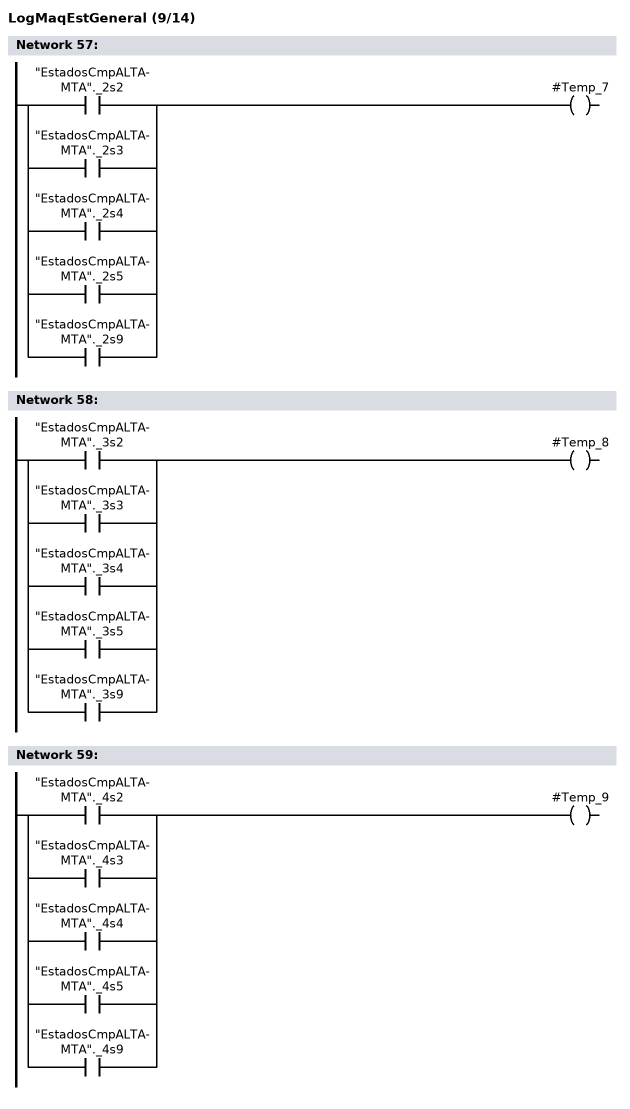
   RUNG wire#powerrail
      Contact( "EstadosCmpALTA-MTA"._2s2 )
      wire#w1
      Coil( #Temp_7 )
   END_RUNG
   RUNG wire#powerrail
      Contact( "EstadosCmpALTA-MTA"._2s3 )
   END_RUNG wire#w1
   RUNG wire#powerrail
      Contact( "EstadosCmpALTA-MTA"._2s4 )
   END_RUNG wire#w1
   RUNG wire#powerrail
      Contact( "EstadosCmpALTA-MTA"._2s5 )
   END_RUNG wire#w1
   RUNG wire#powerrail
      Contact( "EstadosCmpALTA-MTA"._2s9 )
   END_RUNG wire#w1
   // the same network as SCL:
   #Temp_7 := "EstadosCmpALTA-MTA"._2s2 OR "EstadosCmpALTA-MTA"._2s3 OR "EstadosCmpALTA-MTA"._2s4 OR "EstadosCmpALTA-MTA"._2s5 OR "EstadosCmpALTA-MTA"._2s9;
END_REGION

REGION Network 58
   RUNG wire#powerrail
      Contact( "EstadosCmpALTA-MTA"._3s2 )
      wire#w1
      Coil( #Temp_8 )
   END_RUNG
   RUNG wire#powerrail
      Contact( "EstadosCmpALTA-MTA"._3s3 )
   END_RUNG wire#w1
   RUNG wire#powerrail
      Contact( "EstadosCmpALTA-MTA"._3s4 )
   END_RUNG wire#w1
   RUNG wire#powerrail
      Contact( "EstadosCmpALTA-MTA"._3s5 )
   END_RUNG wire#w1
   RUNG wire#powerrail
      Contact( "EstadosCmpALTA-MTA"._3s9 )
   END_RUNG wire#w1
   // the same network as SCL:
   #Temp_8 := "EstadosCmpALTA-MTA"._3s2 OR "EstadosCmpALTA-MTA"._3s3 OR "EstadosCmpALTA-MTA"._3s4 OR "EstadosCmpALTA-MTA"._3s5 OR "EstadosCmpALTA-MTA"._3s9;
END_REGION

REGION Network 59
   RUNG wire#powerrail
      Contact( "EstadosCmpALTA-MTA"._4s2 )
      wire#w1
      Coil( #Temp_9 )
   END_RUNG
   RUNG wire#powerrail
      Contact( "EstadosCmpALTA-MTA"._4s3 )
   END_RUNG wire#w1
   RUNG wire#powerrail
      Contact( "EstadosCmpALTA-MTA"._4s4 )
   END_RUNG wire#w1
   RUNG wire#powerrail
      Contact( "EstadosCmpALTA-MTA"._4s5 )
   END_RUNG wire#w1
   RUNG wire#powerrail
      Contact( "EstadosCmpALTA-MTA"._4s9 )
   END_RUNG wire#w1
   // the same network as SCL:
   #Temp_9 := "EstadosCmpALTA-MTA"._4s2 OR "EstadosCmpALTA-MTA"._4s3 OR "EstadosCmpALTA-MTA"._4s4 OR "EstadosCmpALTA-MTA"._4s5 OR "EstadosCmpALTA-MTA"._4s9;
END_REGION

REGION Network 60
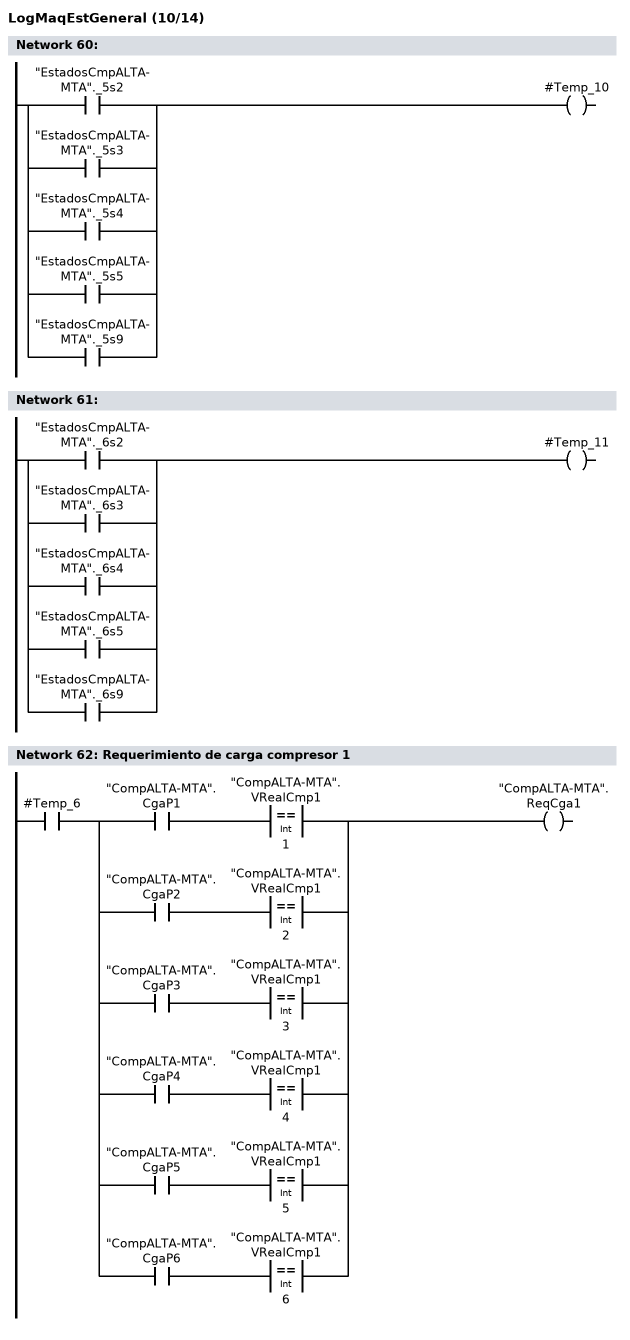
   RUNG wire#powerrail
      Contact( "EstadosCmpALTA-MTA"._5s2 )
      wire#w1
      Coil( #Temp_10 )
   END_RUNG
   RUNG wire#powerrail
      Contact( "EstadosCmpALTA-MTA"._5s3 )
   END_RUNG wire#w1
   RUNG wire#powerrail
      Contact( "EstadosCmpALTA-MTA"._5s4 )
   END_RUNG wire#w1
   RUNG wire#powerrail
      Contact( "EstadosCmpALTA-MTA"._5s5 )
   END_RUNG wire#w1
   RUNG wire#powerrail
      Contact( "EstadosCmpALTA-MTA"._5s9 )
   END_RUNG wire#w1
   // the same network as SCL:
   #Temp_10 := "EstadosCmpALTA-MTA"._5s2 OR "EstadosCmpALTA-MTA"._5s3 OR "EstadosCmpALTA-MTA"._5s4 OR "EstadosCmpALTA-MTA"._5s5 OR "EstadosCmpALTA-MTA"._5s9;
END_REGION

REGION Network 61
   RUNG wire#powerrail
      Contact( "EstadosCmpALTA-MTA"._6s2 )
      wire#w1
      Coil( #Temp_11 )
   END_RUNG
   RUNG wire#powerrail
      Contact( "EstadosCmpALTA-MTA"._6s3 )
   END_RUNG wire#w1
   RUNG wire#powerrail
      Contact( "EstadosCmpALTA-MTA"._6s4 )
   END_RUNG wire#w1
   RUNG wire#powerrail
      Contact( "EstadosCmpALTA-MTA"._6s5 )
   END_RUNG wire#w1
   RUNG wire#powerrail
      Contact( "EstadosCmpALTA-MTA"._6s9 )
   END_RUNG wire#w1
   // the same network as SCL:
   #Temp_11 := "EstadosCmpALTA-MTA"._6s2 OR "EstadosCmpALTA-MTA"._6s3 OR "EstadosCmpALTA-MTA"._6s4 OR "EstadosCmpALTA-MTA"._6s5 OR "EstadosCmpALTA-MTA"._6s9;
END_REGION

REGION Network 62: Requerimiento de carga compresor 1
   RUNG wire#powerrail
      Contact( #Temp_6 )
      wire#w1
      Contact( "CompALTA-MTA".CgaP1 )
      { S7_Templates := "SrcType := Int" } EQ_Contact(in1 := "CompALTA-MTA".VRealCmp1, in2 := 1)
      wire#w2
      Coil( "CompALTA-MTA".ReqCga1 )
   END_RUNG
   RUNG wire#w1
      Contact( "CompALTA-MTA".CgaP2 )
      { S7_Templates := "SrcType := Int" } EQ_Contact(in1 := "CompALTA-MTA".VRealCmp1, in2 := 2)
   END_RUNG wire#w2
   RUNG wire#w1
      Contact( "CompALTA-MTA".CgaP3 )
      { S7_Templates := "SrcType := Int" } EQ_Contact(in1 := "CompALTA-MTA".VRealCmp1, in2 := 3)
   END_RUNG wire#w2
   RUNG wire#w1
      Contact( "CompALTA-MTA".CgaP4 )
      { S7_Templates := "SrcType := Int" } EQ_Contact(in1 := "CompALTA-MTA".VRealCmp1, in2 := 4)
   END_RUNG wire#w2
   RUNG wire#w1
      Contact( "CompALTA-MTA".CgaP5 )
      { S7_Templates := "SrcType := Int" } EQ_Contact(in1 := "CompALTA-MTA".VRealCmp1, in2 := 5)
   END_RUNG wire#w2
   RUNG wire#w1
      Contact( "CompALTA-MTA".CgaP6 )
      { S7_Templates := "SrcType := Int" } EQ_Contact(in1 := "CompALTA-MTA".VRealCmp1, in2 := 6)
   END_RUNG wire#w2
   // the same network as SCL:
   "CompALTA-MTA".ReqCga1 := #Temp_6 AND (("CompALTA-MTA".CgaP1 AND ("CompALTA-MTA".VRealCmp1 = 1)) OR ("CompALTA-MTA".CgaP2 AND ("CompALTA-MTA".VRealCmp1 = 2)) OR ("CompALTA-MTA".CgaP3 AND ("CompALTA-MTA".VRealCmp1 = 3)) OR ("CompALTA-MTA".CgaP4 AND ("CompALTA-MTA".VRealCmp1 = 4)) OR ("CompALTA-MTA".CgaP5 AND ("CompALTA-MTA".VRealCmp1 = 5)) OR ("CompALTA-MTA".CgaP6 AND ("CompALTA-MTA".VRealCmp1 = 6)));
END_REGION

REGION Network 63: Requerimiento de carga compresor 2
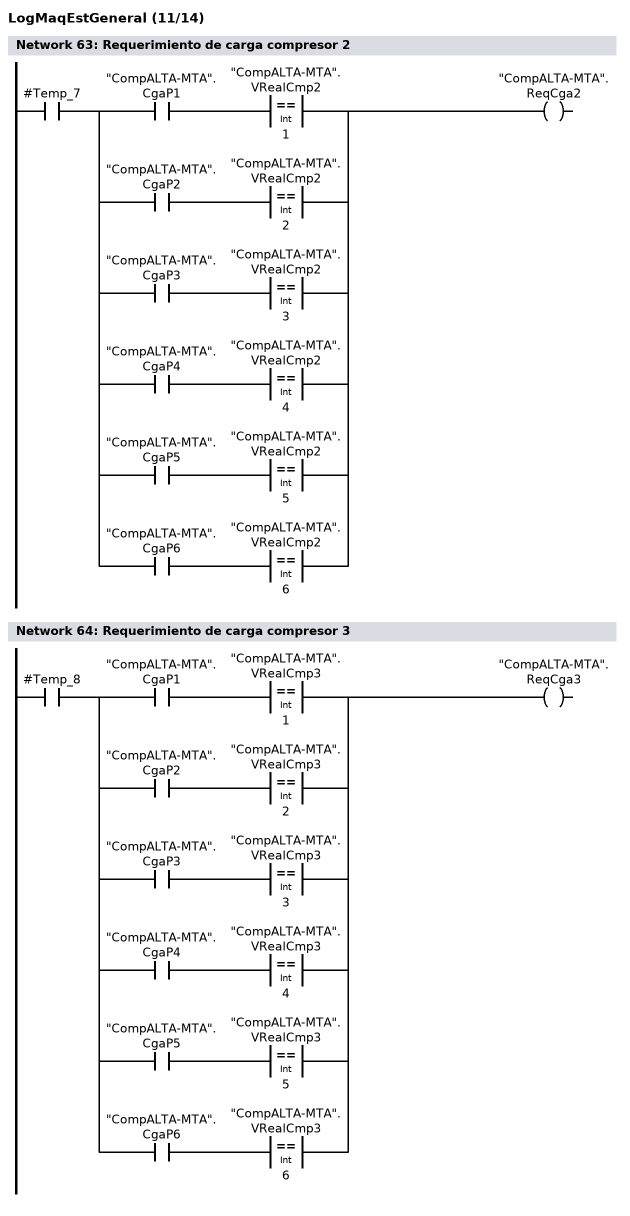
   RUNG wire#powerrail
      Contact( #Temp_7 )
      wire#w1
      Contact( "CompALTA-MTA".CgaP1 )
      { S7_Templates := "SrcType := Int" } EQ_Contact(in1 := "CompALTA-MTA".VRealCmp2, in2 := 1)
      wire#w2
      Coil( "CompALTA-MTA".ReqCga2 )
   END_RUNG
   RUNG wire#w1
      Contact( "CompALTA-MTA".CgaP2 )
      { S7_Templates := "SrcType := Int" } EQ_Contact(in1 := "CompALTA-MTA".VRealCmp2, in2 := 2)
   END_RUNG wire#w2
   RUNG wire#w1
      Contact( "CompALTA-MTA".CgaP3 )
      { S7_Templates := "SrcType := Int" } EQ_Contact(in1 := "CompALTA-MTA".VRealCmp2, in2 := 3)
   END_RUNG wire#w2
   RUNG wire#w1
      Contact( "CompALTA-MTA".CgaP4 )
      { S7_Templates := "SrcType := Int" } EQ_Contact(in1 := "CompALTA-MTA".VRealCmp2, in2 := 4)
   END_RUNG wire#w2
   RUNG wire#w1
      Contact( "CompALTA-MTA".CgaP5 )
      { S7_Templates := "SrcType := Int" } EQ_Contact(in1 := "CompALTA-MTA".VRealCmp2, in2 := 5)
   END_RUNG wire#w2
   RUNG wire#w1
      Contact( "CompALTA-MTA".CgaP6 )
      { S7_Templates := "SrcType := Int" } EQ_Contact(in1 := "CompALTA-MTA".VRealCmp2, in2 := 6)
   END_RUNG wire#w2
   // the same network as SCL:
   "CompALTA-MTA".ReqCga2 := #Temp_7 AND (("CompALTA-MTA".CgaP1 AND ("CompALTA-MTA".VRealCmp2 = 1)) OR ("CompALTA-MTA".CgaP2 AND ("CompALTA-MTA".VRealCmp2 = 2)) OR ("CompALTA-MTA".CgaP3 AND ("CompALTA-MTA".VRealCmp2 = 3)) OR ("CompALTA-MTA".CgaP4 AND ("CompALTA-MTA".VRealCmp2 = 4)) OR ("CompALTA-MTA".CgaP5 AND ("CompALTA-MTA".VRealCmp2 = 5)) OR ("CompALTA-MTA".CgaP6 AND ("CompALTA-MTA".VRealCmp2 = 6)));
END_REGION

REGION Network 64: Requerimiento de carga compresor 3
   RUNG wire#powerrail
      Contact( #Temp_8 )
      wire#w1
      Contact( "CompALTA-MTA".CgaP1 )
      { S7_Templates := "SrcType := Int" } EQ_Contact(in1 := "CompALTA-MTA".VRealCmp3, in2 := 1)
      wire#w2
      Coil( "CompALTA-MTA".ReqCga3 )
   END_RUNG
   RUNG wire#w1
      Contact( "CompALTA-MTA".CgaP2 )
      { S7_Templates := "SrcType := Int" } EQ_Contact(in1 := "CompALTA-MTA".VRealCmp3, in2 := 2)
   END_RUNG wire#w2
   RUNG wire#w1
      Contact( "CompALTA-MTA".CgaP3 )
      { S7_Templates := "SrcType := Int" } EQ_Contact(in1 := "CompALTA-MTA".VRealCmp3, in2 := 3)
   END_RUNG wire#w2
   RUNG wire#w1
      Contact( "CompALTA-MTA".CgaP4 )
      { S7_Templates := "SrcType := Int" } EQ_Contact(in1 := "CompALTA-MTA".VRealCmp3, in2 := 4)
   END_RUNG wire#w2
   RUNG wire#w1
      Contact( "CompALTA-MTA".CgaP5 )
      { S7_Templates := "SrcType := Int" } EQ_Contact(in1 := "CompALTA-MTA".VRealCmp3, in2 := 5)
   END_RUNG wire#w2
   RUNG wire#w1
      Contact( "CompALTA-MTA".CgaP6 )
      { S7_Templates := "SrcType := Int" } EQ_Contact(in1 := "CompALTA-MTA".VRealCmp3, in2 := 6)
   END_RUNG wire#w2
   // the same network as SCL:
   "CompALTA-MTA".ReqCga3 := #Temp_8 AND (("CompALTA-MTA".CgaP1 AND ("CompALTA-MTA".VRealCmp3 = 1)) OR ("CompALTA-MTA".CgaP2 AND ("CompALTA-MTA".VRealCmp3 = 2)) OR ("CompALTA-MTA".CgaP3 AND ("CompALTA-MTA".VRealCmp3 = 3)) OR ("CompALTA-MTA".CgaP4 AND ("CompALTA-MTA".VRealCmp3 = 4)) OR ("CompALTA-MTA".CgaP5 AND ("CompALTA-MTA".VRealCmp3 = 5)) OR ("CompALTA-MTA".CgaP6 AND ("CompALTA-MTA".VRealCmp3 = 6)));
END_REGION

REGION Network 65: Requerimiento de carga compresor 4
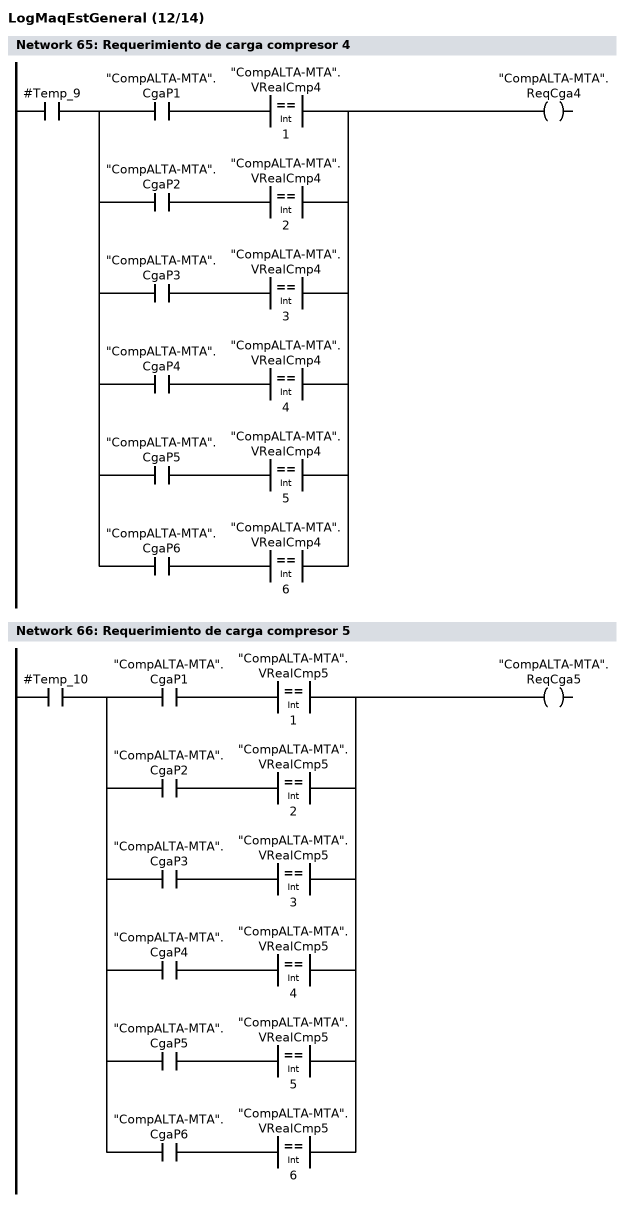
   RUNG wire#powerrail
      Contact( #Temp_9 )
      wire#w1
      Contact( "CompALTA-MTA".CgaP1 )
      { S7_Templates := "SrcType := Int" } EQ_Contact(in1 := "CompALTA-MTA".VRealCmp4, in2 := 1)
      wire#w2
      Coil( "CompALTA-MTA".ReqCga4 )
   END_RUNG
   RUNG wire#w1
      Contact( "CompALTA-MTA".CgaP2 )
      { S7_Templates := "SrcType := Int" } EQ_Contact(in1 := "CompALTA-MTA".VRealCmp4, in2 := 2)
   END_RUNG wire#w2
   RUNG wire#w1
      Contact( "CompALTA-MTA".CgaP3 )
      { S7_Templates := "SrcType := Int" } EQ_Contact(in1 := "CompALTA-MTA".VRealCmp4, in2 := 3)
   END_RUNG wire#w2
   RUNG wire#w1
      Contact( "CompALTA-MTA".CgaP4 )
      { S7_Templates := "SrcType := Int" } EQ_Contact(in1 := "CompALTA-MTA".VRealCmp4, in2 := 4)
   END_RUNG wire#w2
   RUNG wire#w1
      Contact( "CompALTA-MTA".CgaP5 )
      { S7_Templates := "SrcType := Int" } EQ_Contact(in1 := "CompALTA-MTA".VRealCmp4, in2 := 5)
   END_RUNG wire#w2
   RUNG wire#w1
      Contact( "CompALTA-MTA".CgaP6 )
      { S7_Templates := "SrcType := Int" } EQ_Contact(in1 := "CompALTA-MTA".VRealCmp4, in2 := 6)
   END_RUNG wire#w2
   // the same network as SCL:
   "CompALTA-MTA".ReqCga4 := #Temp_9 AND (("CompALTA-MTA".CgaP1 AND ("CompALTA-MTA".VRealCmp4 = 1)) OR ("CompALTA-MTA".CgaP2 AND ("CompALTA-MTA".VRealCmp4 = 2)) OR ("CompALTA-MTA".CgaP3 AND ("CompALTA-MTA".VRealCmp4 = 3)) OR ("CompALTA-MTA".CgaP4 AND ("CompALTA-MTA".VRealCmp4 = 4)) OR ("CompALTA-MTA".CgaP5 AND ("CompALTA-MTA".VRealCmp4 = 5)) OR ("CompALTA-MTA".CgaP6 AND ("CompALTA-MTA".VRealCmp4 = 6)));
END_REGION

REGION Network 66: Requerimiento de carga compresor 5
   RUNG wire#powerrail
      Contact( #Temp_10 )
      wire#w1
      Contact( "CompALTA-MTA".CgaP1 )
      { S7_Templates := "SrcType := Int" } EQ_Contact(in1 := "CompALTA-MTA".VRealCmp5, in2 := 1)
      wire#w2
      Coil( "CompALTA-MTA".ReqCga5 )
   END_RUNG
   RUNG wire#w1
      Contact( "CompALTA-MTA".CgaP2 )
      { S7_Templates := "SrcType := Int" } EQ_Contact(in1 := "CompALTA-MTA".VRealCmp5, in2 := 2)
   END_RUNG wire#w2
   RUNG wire#w1
      Contact( "CompALTA-MTA".CgaP3 )
      { S7_Templates := "SrcType := Int" } EQ_Contact(in1 := "CompALTA-MTA".VRealCmp5, in2 := 3)
   END_RUNG wire#w2
   RUNG wire#w1
      Contact( "CompALTA-MTA".CgaP4 )
      { S7_Templates := "SrcType := Int" } EQ_Contact(in1 := "CompALTA-MTA".VRealCmp5, in2 := 4)
   END_RUNG wire#w2
   RUNG wire#w1
      Contact( "CompALTA-MTA".CgaP5 )
      { S7_Templates := "SrcType := Int" } EQ_Contact(in1 := "CompALTA-MTA".VRealCmp5, in2 := 5)
   END_RUNG wire#w2
   RUNG wire#w1
      Contact( "CompALTA-MTA".CgaP6 )
      { S7_Templates := "SrcType := Int" } EQ_Contact(in1 := "CompALTA-MTA".VRealCmp5, in2 := 6)
   END_RUNG wire#w2
   // the same network as SCL:
   "CompALTA-MTA".ReqCga5 := #Temp_10 AND (("CompALTA-MTA".CgaP1 AND ("CompALTA-MTA".VRealCmp5 = 1)) OR ("CompALTA-MTA".CgaP2 AND ("CompALTA-MTA".VRealCmp5 = 2)) OR ("CompALTA-MTA".CgaP3 AND ("CompALTA-MTA".VRealCmp5 = 3)) OR ("CompALTA-MTA".CgaP4 AND ("CompALTA-MTA".VRealCmp5 = 4)) OR ("CompALTA-MTA".CgaP5 AND ("CompALTA-MTA".VRealCmp5 = 5)) OR ("CompALTA-MTA".CgaP6 AND ("CompALTA-MTA".VRealCmp5 = 6)));
END_REGION

REGION Network 67: Requerimiento de carga compresor 6
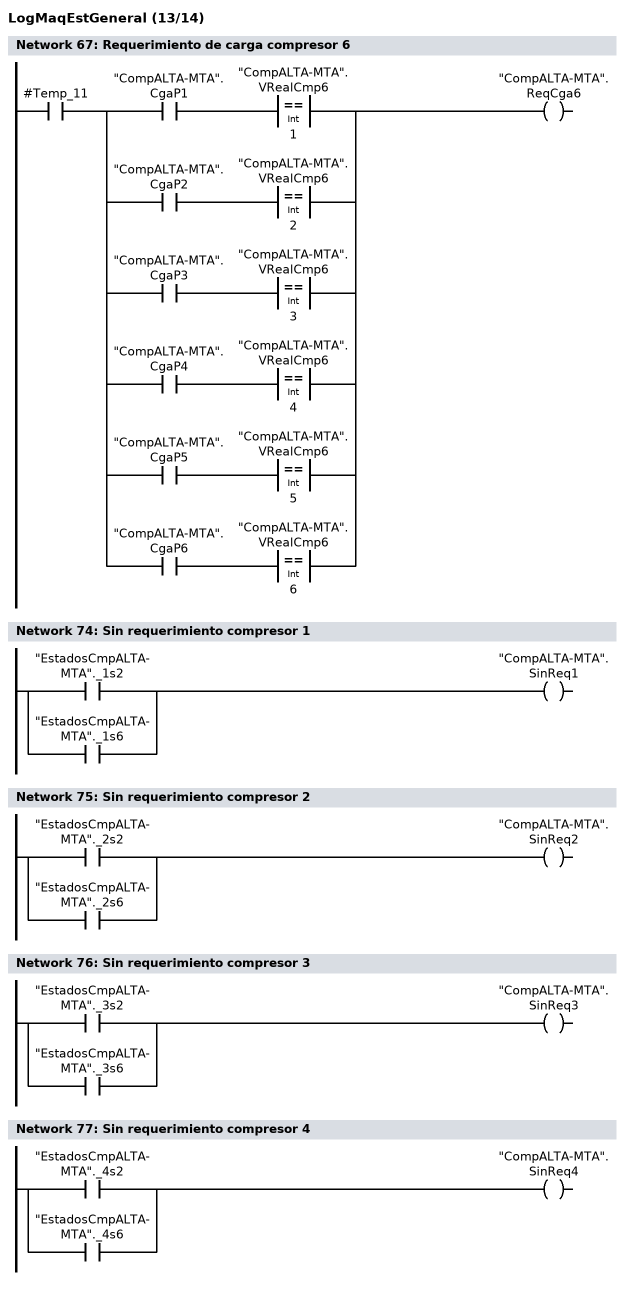
   RUNG wire#powerrail
      Contact( #Temp_11 )
      wire#w1
      Contact( "CompALTA-MTA".CgaP1 )
      { S7_Templates := "SrcType := Int" } EQ_Contact(in1 := "CompALTA-MTA".VRealCmp6, in2 := 1)
      wire#w2
      Coil( "CompALTA-MTA".ReqCga6 )
   END_RUNG
   RUNG wire#w1
      Contact( "CompALTA-MTA".CgaP2 )
      { S7_Templates := "SrcType := Int" } EQ_Contact(in1 := "CompALTA-MTA".VRealCmp6, in2 := 2)
   END_RUNG wire#w2
   RUNG wire#w1
      Contact( "CompALTA-MTA".CgaP3 )
      { S7_Templates := "SrcType := Int" } EQ_Contact(in1 := "CompALTA-MTA".VRealCmp6, in2 := 3)
   END_RUNG wire#w2
   RUNG wire#w1
      Contact( "CompALTA-MTA".CgaP4 )
      { S7_Templates := "SrcType := Int" } EQ_Contact(in1 := "CompALTA-MTA".VRealCmp6, in2 := 4)
   END_RUNG wire#w2
   RUNG wire#w1
      Contact( "CompALTA-MTA".CgaP5 )
      { S7_Templates := "SrcType := Int" } EQ_Contact(in1 := "CompALTA-MTA".VRealCmp6, in2 := 5)
   END_RUNG wire#w2
   RUNG wire#w1
      Contact( "CompALTA-MTA".CgaP6 )
      { S7_Templates := "SrcType := Int" } EQ_Contact(in1 := "CompALTA-MTA".VRealCmp6, in2 := 6)
   END_RUNG wire#w2
   // the same network as SCL:
   "CompALTA-MTA".ReqCga6 := #Temp_11 AND (("CompALTA-MTA".CgaP1 AND ("CompALTA-MTA".VRealCmp6 = 1)) OR ("CompALTA-MTA".CgaP2 AND ("CompALTA-MTA".VRealCmp6 = 2)) OR ("CompALTA-MTA".CgaP3 AND ("CompALTA-MTA".VRealCmp6 = 3)) OR ("CompALTA-MTA".CgaP4 AND ("CompALTA-MTA".VRealCmp6 = 4)) OR ("CompALTA-MTA".CgaP5 AND ("CompALTA-MTA".VRealCmp6 = 5)) OR ("CompALTA-MTA".CgaP6 AND ("CompALTA-MTA".VRealCmp6 = 6)));
END_REGION

REGION Network 68 (STL)
         A(;
         L     "DB-PrioridadesCmpAlta".Vcmp1;
         L     1;
         ==R;
         );
         AN    "DB-CompAltaDatos".Aut1;
         O;
         A(;
         L     "DB-PrioridadesCmpAlta".Vcmp2;
         L     1;
         ==R;
         );
         AN    "DB-CompAltaDatos".Aut2;
         O;
         A(;
         L     "DB-PrioridadesCmpAlta".Vcmp3;
         L     1;
         ==R;
         );
         AN    "DB-CompAltaDatos".Aut3;
         O;
         A(;
         L     "DB-PrioridadesCmpAlta".Vcmp4;
         L     1;
         ==R;
         );
         AN    "DB-CompAltaDatos".Aut4;
         O;
         A(;
         L     "DB-PrioridadesCmpAlta".Vcmp5;
         L     1;
         ==R;
         );
         AN    "DB-CompAltaDatos".Aut5;
         O;
         A(;
         L     "DB-PrioridadesCmpAlta".Vcmp6;
         L     1;
         ==R;
         );
         AN    "DB-CompAltaDatos".Aut6;
         =     "CompALTA-MTA".ManP1;
END_REGION

REGION Network 69 (STL)
         A(;
         L     "DB-PrioridadesCmpAlta".Vcmp1;
         L     2;
         ==R;
         );
         AN    "DB-CompAltaDatos".Aut1;
         O;
         A(;
         L     "DB-PrioridadesCmpAlta".Vcmp2;
         L     2;
         ==R;
         );
         AN    "DB-CompAltaDatos".Aut2;
         O;
         A(;
         L     "DB-PrioridadesCmpAlta".Vcmp3;
         L     2;
         ==R;
         );
         AN    "DB-CompAltaDatos".Aut3;
         O;
         A(;
         L     "DB-PrioridadesCmpAlta".Vcmp4;
         L     2;
         ==R;
         );
         AN    "DB-CompAltaDatos".Aut4;
         O;
         A(;
         L     "DB-PrioridadesCmpAlta".Vcmp5;
         L     2;
         ==R;
         );
         AN    "DB-CompAltaDatos".Aut5;
         A(;
         L     "DB-PrioridadesCmpAlta".Vcmp6;
         L     2;
         ==R;
         );
         AN    "DB-CompAltaDatos".Aut6;
         =     "CompALTA-MTA".ManP2;
END_REGION

REGION Network 70 (STL)
         A(;
         L     "DB-PrioridadesCmpAlta".Vcmp1;
         L     3;
         ==R;
         );
         AN    "DB-CompAltaDatos".Aut1;
         O;
         A(;
         L     "DB-PrioridadesCmpAlta".Vcmp2;
         L     3;
         ==R;
         );
         AN    "DB-CompAltaDatos".Aut2;
         O;
         A(;
         L     "DB-PrioridadesCmpAlta".Vcmp3;
         L     3;
         ==R;
         );
         AN    "DB-CompAltaDatos".Aut3;
         O;
         A(;
         L     "DB-PrioridadesCmpAlta".Vcmp4;
         L     3;
         ==R;
         );
         AN    "DB-CompAltaDatos".Aut4;
         O;
         A(;
         L     "DB-PrioridadesCmpAlta".Vcmp5;
         L     3;
         ==R;
         );
         AN    "DB-CompAltaDatos".Aut5;
         O;
         A(;
         L     "DB-PrioridadesCmpAlta".Vcmp6;
         L     3;
         ==R;
         );
         AN    "DB-CompAltaDatos".Aut6;
         =     "CompALTA-MTA".ManP3;
END_REGION

REGION Network 71 (STL)
         A(;
         L     "DB-PrioridadesCmpAlta".Vcmp1;
         L     4;
         ==R;
         );
         AN    "DB-CompAltaDatos".Aut1;
         O;
         A(;
         L     "DB-PrioridadesCmpAlta".Vcmp2;
         L     4;
         ==R;
         );
         AN    "DB-CompAltaDatos".Aut2;
         O;
         A(;
         L     "DB-PrioridadesCmpAlta".Vcmp3;
         L     4;
         ==R;
         );
         AN    "DB-CompAltaDatos".Aut3;
         O;
         A(;
         L     "DB-PrioridadesCmpAlta".Vcmp4;
         L     4;
         ==R;
         );
         AN    "DB-CompAltaDatos".Aut4;
         O;
         A(;
         L     "DB-PrioridadesCmpAlta".Vcmp5;
         L     4;
         ==R;
         );
         AN    "DB-CompAltaDatos".Aut5;
         O;
         A(;
         L     "DB-PrioridadesCmpAlta".Vcmp6;
         L     4;
         ==R;
         );
         AN    "DB-CompAltaDatos".Aut6;
         =     "CompALTA-MTA".ManP4;
END_REGION

REGION Network 72 (STL)
         A(;
         L     "DB-PrioridadesCmpAlta".Vcmp1;
         L     5;
         ==R;
         );
         AN    "DB-CompAltaDatos".Aut1;
         O;
         A(;
         L     "DB-PrioridadesCmpAlta".Vcmp2;
         L     5;
         ==R;
         );
         AN    "DB-CompAltaDatos".Aut2;
         O;
         A(;
         L     "DB-PrioridadesCmpAlta".Vcmp3;
         L     5;
         ==R;
         );
         AN    "DB-CompAltaDatos".Aut3;
         O;
         A(;
         L     "DB-PrioridadesCmpAlta".Vcmp4;
         L     5;
         ==R;
         );
         AN    "DB-CompAltaDatos".Aut4;
         O;
         A(;
         L     "DB-PrioridadesCmpAlta".Vcmp5;
         L     5;
         ==R;
         );
         AN    "DB-CompAltaDatos".Aut5;
         O;
         A(;
         L     "DB-PrioridadesCmpAlta".Vcmp6;
         L     5;
         ==R;
         );
         AN    "DB-CompAltaDatos".Aut6;
         =     "CompALTA-MTA".ManP5;
END_REGION

REGION Network 73 (STL)
         A(;
         L     "DB-PrioridadesCmpAlta".Vcmp1;
         L     6;
         ==R;
         );
         AN    "DB-CompAltaDatos".Aut1;
         O;
         A(;
         L     "DB-PrioridadesCmpAlta".Vcmp2;
         L     6;
         ==R;
         );
         AN    "DB-CompAltaDatos".Aut2;
         O;
         A(;
         L     "DB-PrioridadesCmpAlta".Vcmp3;
         L     6;
         ==R;
         );
         AN    "DB-CompAltaDatos".Aut3;
         O;
         A(;
         L     "DB-PrioridadesCmpAlta".Vcmp4;
         L     6;
         ==R;
         );
         AN    "DB-CompAltaDatos".Aut4;
         O;
         A(;
         L     "DB-PrioridadesCmpAlta".Vcmp5;
         L     6;
         ==R;
         );
         AN    "DB-CompAltaDatos".Aut5;
         O;
         A(;
         L     "DB-PrioridadesCmpAlta".Vcmp6;
         L     6;
         ==R;
         );
         AN    "DB-CompAltaDatos".Aut6;
         =     "CompALTA-MTA".ManP6;
END_REGION

REGION Network 74: Sin requerimiento compresor 1
   RUNG wire#powerrail
      Contact( "EstadosCmpALTA-MTA"._1s2 )
      wire#w1
      Coil( "CompALTA-MTA".SinReq1 )
   END_RUNG
   RUNG wire#powerrail
      Contact( "EstadosCmpALTA-MTA"._1s6 )
   END_RUNG wire#w1
   // the same network as SCL:
   "CompALTA-MTA".SinReq1 := "EstadosCmpALTA-MTA"._1s2 OR "EstadosCmpALTA-MTA"._1s6;
END_REGION

REGION Network 75: Sin requerimiento compresor 2
   RUNG wire#powerrail
      Contact( "EstadosCmpALTA-MTA"._2s2 )
      wire#w1
      Coil( "CompALTA-MTA".SinReq2 )
   END_RUNG
   RUNG wire#powerrail
      Contact( "EstadosCmpALTA-MTA"._2s6 )
   END_RUNG wire#w1
   // the same network as SCL:
   "CompALTA-MTA".SinReq2 := "EstadosCmpALTA-MTA"._2s2 OR "EstadosCmpALTA-MTA"._2s6;
END_REGION

REGION Network 76: Sin requerimiento compresor 3
   RUNG wire#powerrail
      Contact( "EstadosCmpALTA-MTA"._3s2 )
      wire#w1
      Coil( "CompALTA-MTA".SinReq3 )
   END_RUNG
   RUNG wire#powerrail
      Contact( "EstadosCmpALTA-MTA"._3s6 )
   END_RUNG wire#w1
   // the same network as SCL:
   "CompALTA-MTA".SinReq3 := "EstadosCmpALTA-MTA"._3s2 OR "EstadosCmpALTA-MTA"._3s6;
END_REGION

REGION Network 77: Sin requerimiento compresor 4
   RUNG wire#powerrail
      Contact( "EstadosCmpALTA-MTA"._4s2 )
      wire#w1
      Coil( "CompALTA-MTA".SinReq4 )
   END_RUNG
   RUNG wire#powerrail
      Contact( "EstadosCmpALTA-MTA"._4s6 )
   END_RUNG wire#w1
   // the same network as SCL:
   "CompALTA-MTA".SinReq4 := "EstadosCmpALTA-MTA"._4s2 OR "EstadosCmpALTA-MTA"._4s6;
END_REGION

REGION Network 78: Sin requerimiento compresor 5
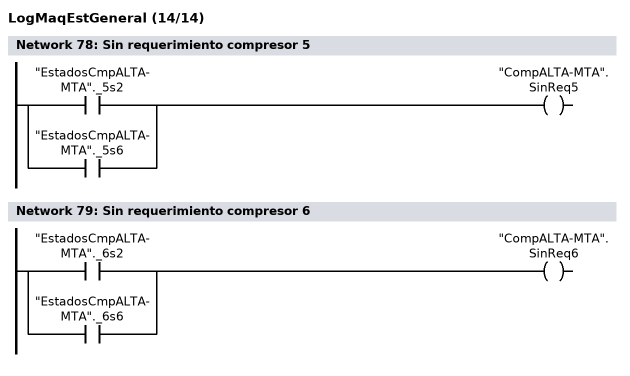
   RUNG wire#powerrail
      Contact( "EstadosCmpALTA-MTA"._5s2 )
      wire#w1
      Coil( "CompALTA-MTA".SinReq5 )
   END_RUNG
   RUNG wire#powerrail
      Contact( "EstadosCmpALTA-MTA"._5s6 )
   END_RUNG wire#w1
   // the same network as SCL:
   "CompALTA-MTA".SinReq5 := "EstadosCmpALTA-MTA"._5s2 OR "EstadosCmpALTA-MTA"._5s6;
END_REGION

REGION Network 79: Sin requerimiento compresor 6
   RUNG wire#powerrail
      Contact( "EstadosCmpALTA-MTA"._6s2 )
      wire#w1
      Coil( "CompALTA-MTA".SinReq6 )
   END_RUNG
   RUNG wire#powerrail
      Contact( "EstadosCmpALTA-MTA"._6s6 )
   END_RUNG wire#w1
   // the same network as SCL:
   "CompALTA-MTA".SinReq6 := "EstadosCmpALTA-MTA"._6s2 OR "EstadosCmpALTA-MTA"._6s6;
END_REGION
END_FUNCTION

FUNCTION "CalcEst1" : Void   // FC36, LAD
{ S7_Optimized_Access := 'FALSE' }
VERSION : 0.1
   VAR_TEMP   // added for the SCL form of the ladder/FBD networks
      _w1 : Bool;
   END_VAR
BEGIN

REGION Network 1
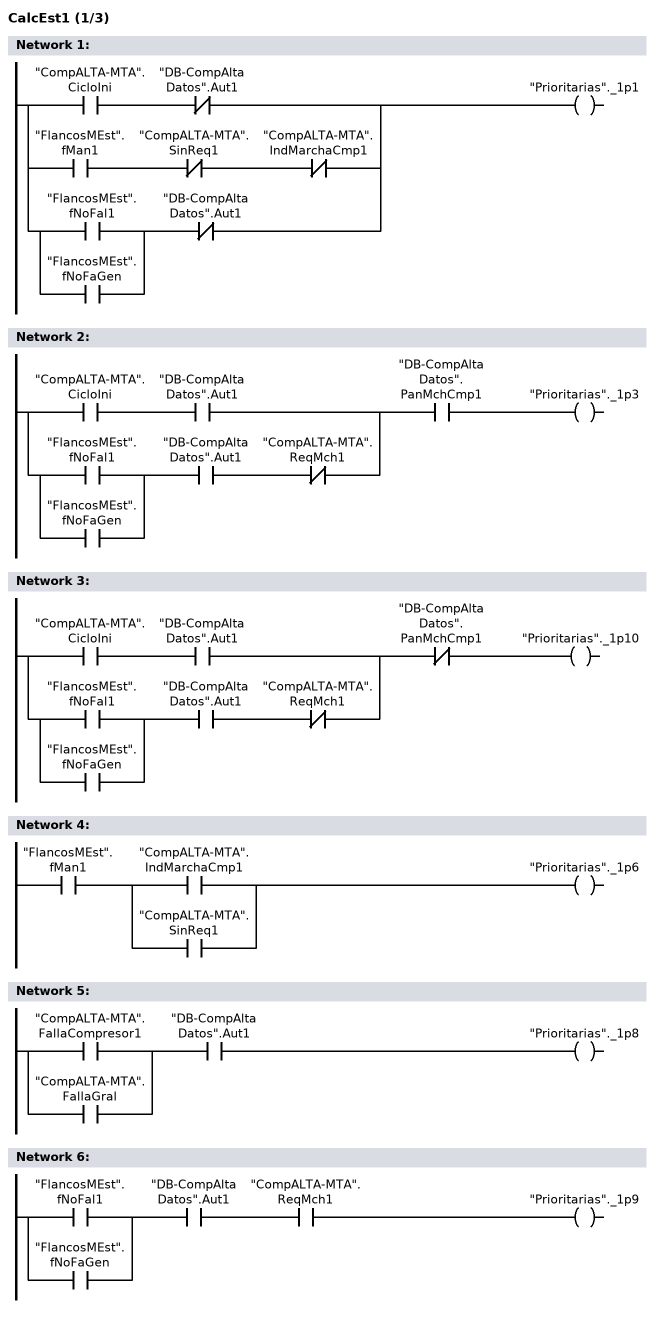
   RUNG wire#powerrail
      Contact( "CompALTA-MTA".CicloIni )
      I_Contact( "DB-CompAltaDatos".Aut1 )
      wire#w1
      Coil( "Prioritarias"._1p1 )
   END_RUNG
   RUNG wire#powerrail
      Contact( "FlancosMEst".fMan1 )
      I_Contact( "CompALTA-MTA".SinReq1 )
      I_Contact( "CompALTA-MTA".IndMarchaCmp1 )
   END_RUNG wire#w1
   RUNG wire#powerrail
      Contact( "FlancosMEst".fNoFal1 )
      wire#w2
      I_Contact( "DB-CompAltaDatos".Aut1 )
   END_RUNG wire#w1
   RUNG wire#powerrail
      Contact( "FlancosMEst".fNoFaGen )
   END_RUNG wire#w2
   // the same network as SCL:
   "Prioritarias"._1p1 := ("CompALTA-MTA".CicloIni AND NOT "DB-CompAltaDatos".Aut1) OR ("FlancosMEst".fMan1 AND NOT "CompALTA-MTA".SinReq1 AND NOT "CompALTA-MTA".IndMarchaCmp1) OR (("FlancosMEst".fNoFal1 OR "FlancosMEst".fNoFaGen) AND NOT "DB-CompAltaDatos".Aut1);
END_REGION

REGION Network 2
   RUNG wire#powerrail
      Contact( "CompALTA-MTA".CicloIni )
      Contact( "DB-CompAltaDatos".Aut1 )
      wire#w1
      Contact( "DB-CompAltaDatos".PanMchCmp1 )
      Coil( "Prioritarias"._1p3 )
   END_RUNG
   RUNG wire#powerrail
      Contact( "FlancosMEst".fNoFal1 )
      wire#w2
      Contact( "DB-CompAltaDatos".Aut1 )
      I_Contact( "CompALTA-MTA".ReqMch1 )
   END_RUNG wire#w1
   RUNG wire#powerrail
      Contact( "FlancosMEst".fNoFaGen )
   END_RUNG wire#w2
   // the same network as SCL:
   "Prioritarias"._1p3 := (("CompALTA-MTA".CicloIni AND "DB-CompAltaDatos".Aut1) OR (("FlancosMEst".fNoFal1 OR "FlancosMEst".fNoFaGen) AND "DB-CompAltaDatos".Aut1 AND NOT "CompALTA-MTA".ReqMch1)) AND "DB-CompAltaDatos".PanMchCmp1;
END_REGION

REGION Network 3
   RUNG wire#powerrail
      Contact( "CompALTA-MTA".CicloIni )
      Contact( "DB-CompAltaDatos".Aut1 )
      wire#w1
      I_Contact( "DB-CompAltaDatos".PanMchCmp1 )
      Coil( "Prioritarias"._1p10 )
   END_RUNG
   RUNG wire#powerrail
      Contact( "FlancosMEst".fNoFal1 )
      wire#w2
      Contact( "DB-CompAltaDatos".Aut1 )
      I_Contact( "CompALTA-MTA".ReqMch1 )
   END_RUNG wire#w1
   RUNG wire#powerrail
      Contact( "FlancosMEst".fNoFaGen )
   END_RUNG wire#w2
   // the same network as SCL:
   "Prioritarias"._1p10 := (("CompALTA-MTA".CicloIni AND "DB-CompAltaDatos".Aut1) OR (("FlancosMEst".fNoFal1 OR "FlancosMEst".fNoFaGen) AND "DB-CompAltaDatos".Aut1 AND NOT "CompALTA-MTA".ReqMch1)) AND NOT "DB-CompAltaDatos".PanMchCmp1;
END_REGION

REGION Network 4
   RUNG wire#powerrail
      Contact( "FlancosMEst".fMan1 )
      wire#w1
      Contact( "CompALTA-MTA".IndMarchaCmp1 )
      wire#w2
      Coil( "Prioritarias"._1p6 )
   END_RUNG
   RUNG wire#w1
      Contact( "CompALTA-MTA".SinReq1 )
   END_RUNG wire#w2
   // the same network as SCL:
   "Prioritarias"._1p6 := "FlancosMEst".fMan1 AND ("CompALTA-MTA".IndMarchaCmp1 OR "CompALTA-MTA".SinReq1);
END_REGION

REGION Network 5
   RUNG wire#powerrail
      Contact( "CompALTA-MTA".FallaCompresor1 )
      wire#w1
      Contact( "DB-CompAltaDatos".Aut1 )
      Coil( "Prioritarias"._1p8 )
   END_RUNG
   RUNG wire#powerrail
      Contact( "CompALTA-MTA".FallaGral )
   END_RUNG wire#w1
   // the same network as SCL:
   "Prioritarias"._1p8 := ("CompALTA-MTA".FallaCompresor1 OR "CompALTA-MTA".FallaGral) AND "DB-CompAltaDatos".Aut1;
END_REGION

REGION Network 6
   RUNG wire#powerrail
      Contact( "FlancosMEst".fNoFal1 )
      wire#w1
      Contact( "DB-CompAltaDatos".Aut1 )
      Contact( "CompALTA-MTA".ReqMch1 )
      Coil( "Prioritarias"._1p9 )
   END_RUNG
   RUNG wire#powerrail
      Contact( "FlancosMEst".fNoFaGen )
   END_RUNG wire#w1
   // the same network as SCL:
   "Prioritarias"._1p9 := ("FlancosMEst".fNoFal1 OR "FlancosMEst".fNoFaGen) AND "DB-CompAltaDatos".Aut1 AND "CompALTA-MTA".ReqMch1;
END_REGION

REGION Network 7
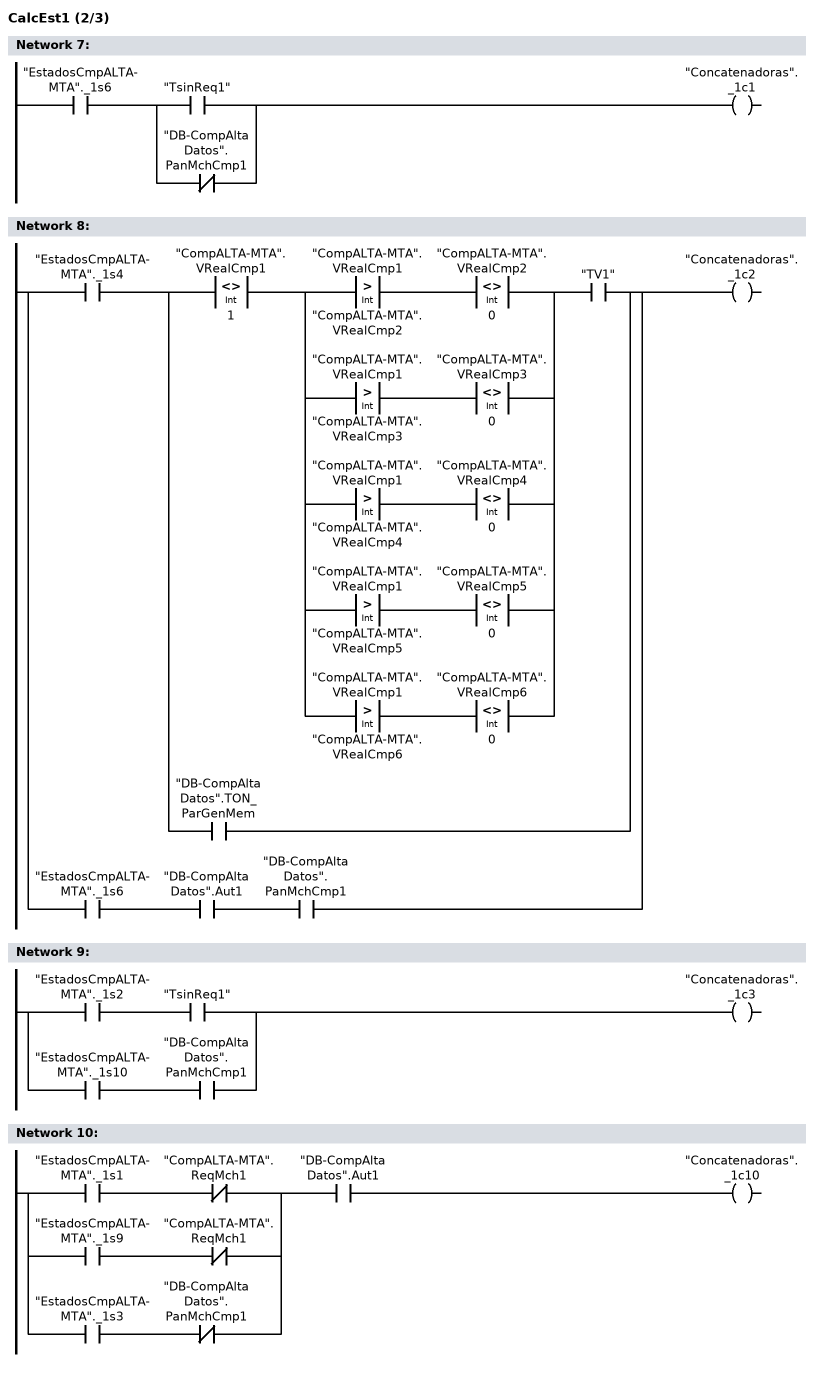
   RUNG wire#powerrail
      Contact( "EstadosCmpALTA-MTA"._1s6 )
      wire#w1
      Contact( "TsinReq1" )
      wire#w2
      Coil( "Concatenadoras"._1c1 )
   END_RUNG
   RUNG wire#w1
      I_Contact( "DB-CompAltaDatos".PanMchCmp1 )
   END_RUNG wire#w2
   // the same network as SCL:
   "Concatenadoras"._1c1 := "EstadosCmpALTA-MTA"._1s6 AND ("TsinReq1" OR NOT "DB-CompAltaDatos".PanMchCmp1);
END_REGION

REGION Network 8
   RUNG wire#powerrail
      Contact( "EstadosCmpALTA-MTA"._1s4 )
      wire#w1
      { S7_Templates := "SrcType := Int" } NE_Contact(in1 := "CompALTA-MTA".VRealCmp1, in2 := 1)
      wire#w2
      { S7_Templates := "SrcType := Int" } GT_Contact(in1 := "CompALTA-MTA".VRealCmp1, in2 := "CompALTA-MTA".VRealCmp2)
      { S7_Templates := "SrcType := Int" } NE_Contact(in1 := "CompALTA-MTA".VRealCmp2, in2 := 0)
      wire#w3
      Contact( "TV1" )
      wire#w4
      Coil( "Concatenadoras"._1c2 )
   END_RUNG
   RUNG wire#w2
      { S7_Templates := "SrcType := Int" } GT_Contact(in1 := "CompALTA-MTA".VRealCmp1, in2 := "CompALTA-MTA".VRealCmp3)
      { S7_Templates := "SrcType := Int" } NE_Contact(in1 := "CompALTA-MTA".VRealCmp3, in2 := 0)
   END_RUNG wire#w3
   RUNG wire#w2
      { S7_Templates := "SrcType := Int" } GT_Contact(in1 := "CompALTA-MTA".VRealCmp1, in2 := "CompALTA-MTA".VRealCmp4)
      { S7_Templates := "SrcType := Int" } NE_Contact(in1 := "CompALTA-MTA".VRealCmp4, in2 := 0)
   END_RUNG wire#w3
   RUNG wire#w2
      { S7_Templates := "SrcType := Int" } GT_Contact(in1 := "CompALTA-MTA".VRealCmp1, in2 := "CompALTA-MTA".VRealCmp5)
      { S7_Templates := "SrcType := Int" } NE_Contact(in1 := "CompALTA-MTA".VRealCmp5, in2 := 0)
   END_RUNG wire#w3
   RUNG wire#w2
      { S7_Templates := "SrcType := Int" } GT_Contact(in1 := "CompALTA-MTA".VRealCmp1, in2 := "CompALTA-MTA".VRealCmp6)
      { S7_Templates := "SrcType := Int" } NE_Contact(in1 := "CompALTA-MTA".VRealCmp6, in2 := 0)
   END_RUNG wire#w3
   RUNG wire#w1
      Contact( "DB-CompAltaDatos".TON_ParGenMem )
   END_RUNG wire#w4
   RUNG wire#powerrail
      Contact( "EstadosCmpALTA-MTA"._1s6 )
      Contact( "DB-CompAltaDatos".Aut1 )
      Contact( "DB-CompAltaDatos".PanMchCmp1 )
   END_RUNG wire#w4
   // the same network as SCL:
   "Concatenadoras"._1c2 := ("EstadosCmpALTA-MTA"._1s4 AND ((("CompALTA-MTA".VRealCmp1 <> 1) AND ((("CompALTA-MTA".VRealCmp1 > "CompALTA-MTA".VRealCmp2) AND ("CompALTA-MTA".VRealCmp2 <> 0)) OR (("CompALTA-MTA".VRealCmp1 > "CompALTA-MTA".VRealCmp3) AND ("CompALTA-MTA".VRealCmp3 <> 0)) OR (("CompALTA-MTA".VRealCmp1 > "CompALTA-MTA".VRealCmp4) AND ("CompALTA-MTA".VRealCmp4 <> 0)) OR (("CompALTA-MTA".VRealCmp1 > "CompALTA-MTA".VRealCmp5) AND ("CompALTA-MTA".VRealCmp5 <> 0)) OR (("CompALTA-MTA".VRealCmp1 > "CompALTA-MTA".VRealCmp6) AND ("CompALTA-MTA".VRealCmp6 <> 0))) AND "TV1") OR "DB-CompAltaDatos".TON_ParGenMem)) OR ("EstadosCmpALTA-MTA"._1s6 AND "DB-CompAltaDatos".Aut1 AND "DB-CompAltaDatos".PanMchCmp1);
END_REGION

REGION Network 9
   RUNG wire#powerrail
      Contact( "EstadosCmpALTA-MTA"._1s2 )
      Contact( "TsinReq1" )
      wire#w1
      Coil( "Concatenadoras"._1c3 )
   END_RUNG
   RUNG wire#powerrail
      Contact( "EstadosCmpALTA-MTA"._1s10 )
      Contact( "DB-CompAltaDatos".PanMchCmp1 )
   END_RUNG wire#w1
   // the same network as SCL:
   "Concatenadoras"._1c3 := ("EstadosCmpALTA-MTA"._1s2 AND "TsinReq1") OR ("EstadosCmpALTA-MTA"._1s10 AND "DB-CompAltaDatos".PanMchCmp1);
END_REGION
